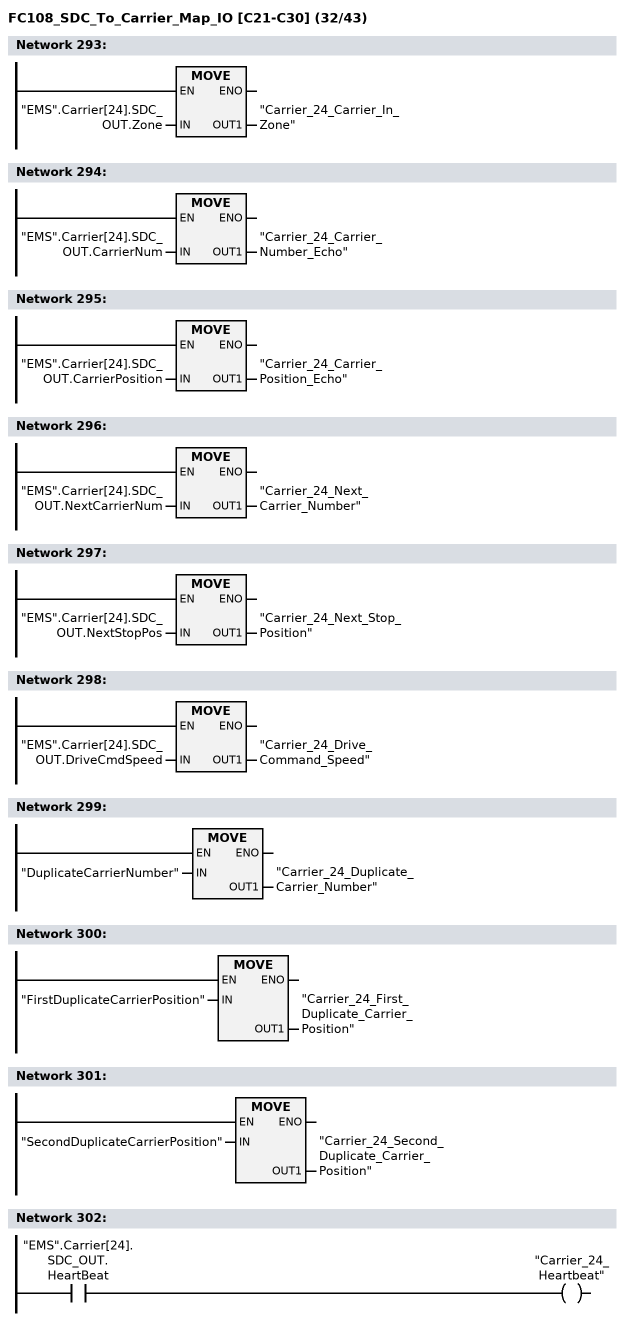
   RUNG wire#powerrail
      Move(in := "EMS".Carrier[24].SDC_OUT.Zone, out1 => "Carrier_24_Carrier_In_Zone")
   END_RUNG
   // the same network as SCL:
   "Carrier_24_Carrier_In_Zone" := "EMS".Carrier[24].SDC_OUT.Zone;
END_REGION

REGION Network 294
   RUNG wire#powerrail
      Move(in := "EMS".Carrier[24].SDC_OUT.CarrierNum, out1 => "Carrier_24_Carrier_Number_Echo")
   END_RUNG
   // the same network as SCL:
   "Carrier_24_Carrier_Number_Echo" := "EMS".Carrier[24].SDC_OUT.CarrierNum;
END_REGION

REGION Network 295
   RUNG wire#powerrail
      Move(in := "EMS".Carrier[24].SDC_OUT.CarrierPosition, out1 => "Carrier_24_Carrier_Position_Echo")
   END_RUNG
   // the same network as SCL:
   "Carrier_24_Carrier_Position_Echo" := "EMS".Carrier[24].SDC_OUT.CarrierPosition;
END_REGION

REGION Network 296
   RUNG wire#powerrail
      Move(in := "EMS".Carrier[24].SDC_OUT.NextCarrierNum, out1 => "Carrier_24_Next_Carrier_Number")
   END_RUNG
   // the same network as SCL:
   "Carrier_24_Next_Carrier_Number" := "EMS".Carrier[24].SDC_OUT.NextCarrierNum;
END_REGION

REGION Network 297
   RUNG wire#powerrail
      Move(in := "EMS".Carrier[24].SDC_OUT.NextStopPos, out1 => "Carrier_24_Next_Stop_Position")
   END_RUNG
   // the same network as SCL:
   "Carrier_24_Next_Stop_Position" := "EMS".Carrier[24].SDC_OUT.NextStopPos;
END_REGION

REGION Network 298
   RUNG wire#powerrail
      Move(in := "EMS".Carrier[24].SDC_OUT.DriveCmdSpeed, out1 => "Carrier_24_Drive_Command_Speed")
   END_RUNG
   // the same network as SCL:
   "Carrier_24_Drive_Command_Speed" := "EMS".Carrier[24].SDC_OUT.DriveCmdSpeed;
END_REGION

REGION Network 299
   RUNG wire#powerrail
      Move(in := "DuplicateCarrierNumber", out1 => "Carrier_24_Duplicate_Carrier_Number")
   END_RUNG
   // the same network as SCL:
   "Carrier_24_Duplicate_Carrier_Number" := "DuplicateCarrierNumber";
END_REGION

REGION Network 300
   RUNG wire#powerrail
      Move(in := "FirstDuplicateCarrierPosition", out1 => "Carrier_24_First_Duplicate_Carrier_Position")
   END_RUNG
   // the same network as SCL:
   "Carrier_24_First_Duplicate_Carrier_Position" := "FirstDuplicateCarrierPosition";
END_REGION

REGION Network 301
   RUNG wire#powerrail
      Move(in := "SecondDuplicateCarrierPosition", out1 => "Carrier_24_Second_Duplicate_Carrier_Position")
   END_RUNG
   // the same network as SCL:
   "Carrier_24_Second_Duplicate_Carrier_Position" := "SecondDuplicateCarrierPosition";
END_REGION

REGION Network 302
   RUNG wire#powerrail
      Contact( "EMS".Carrier[24].SDC_OUT.HeartBeat )
      Coil( "Carrier_24_Heartbeat" )
   END_RUNG
   // the same network as SCL:
   "Carrier_24_Heartbeat" := "EMS".Carrier[24].SDC_OUT.HeartBeat;
END_REGION

REGION Network 303
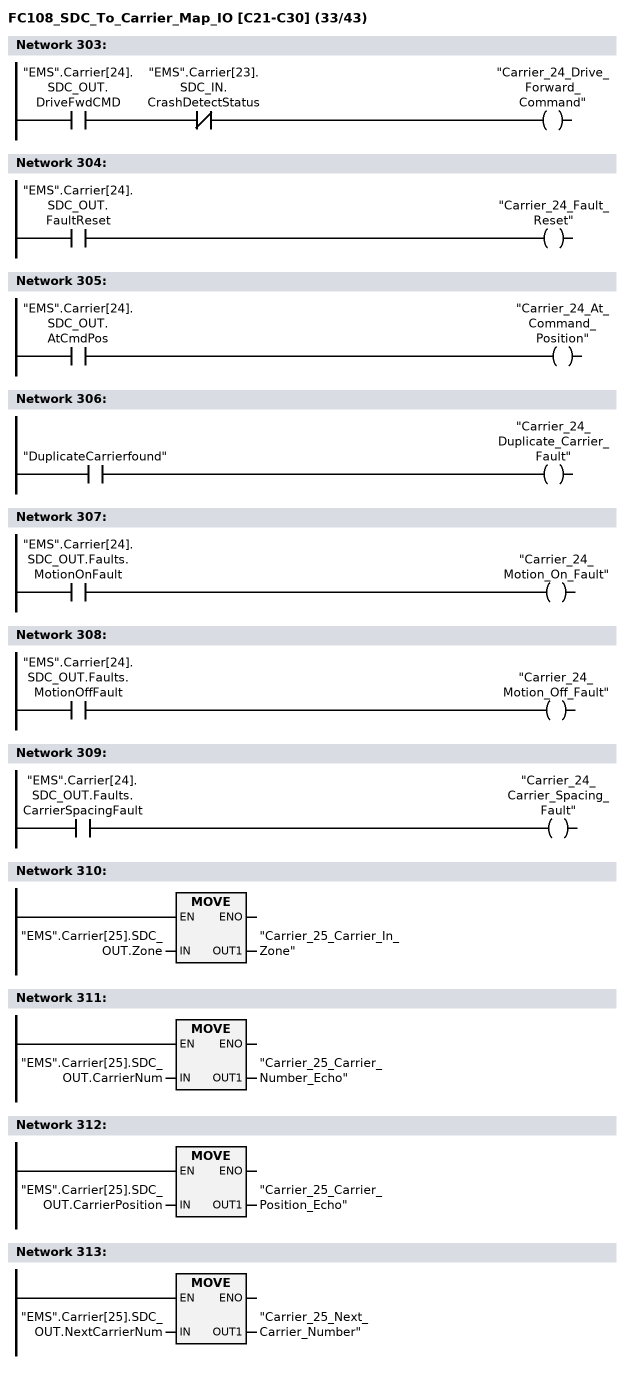
   RUNG wire#powerrail
      Contact( "EMS".Carrier[24].SDC_OUT.DriveFwdCMD )
      I_Contact( "EMS".Carrier[23].SDC_IN.CrashDetectStatus )
      Coil( "Carrier_24_Drive_Forward_Command" )
   END_RUNG
   // the same network as SCL:
   "Carrier_24_Drive_Forward_Command" := "EMS".Carrier[24].SDC_OUT.DriveFwdCMD AND NOT "EMS".Carrier[23].SDC_IN.CrashDetectStatus;
END_REGION

REGION Network 304
   RUNG wire#powerrail
      Contact( "EMS".Carrier[24].SDC_OUT.FaultReset )
      Coil( "Carrier_24_Fault_Reset" )
   END_RUNG
   // the same network as SCL:
   "Carrier_24_Fault_Reset" := "EMS".Carrier[24].SDC_OUT.FaultReset;
END_REGION

REGION Network 305
   RUNG wire#powerrail
      Contact( "EMS".Carrier[24].SDC_OUT.AtCmdPos )
      Coil( "Carrier_24_At_Command_Position" )
   END_RUNG
   // the same network as SCL:
   "Carrier_24_At_Command_Position" := "EMS".Carrier[24].SDC_OUT.AtCmdPos;
END_REGION

REGION Network 306
   RUNG wire#powerrail
      Contact( "DuplicateCarrierfound" )
      Coil( "Carrier_24_Duplicate_Carrier_Fault" )
   END_RUNG
   // the same network as SCL:
   "Carrier_24_Duplicate_Carrier_Fault" := "DuplicateCarrierfound";
END_REGION

REGION Network 307
   RUNG wire#powerrail
      Contact( "EMS".Carrier[24].SDC_OUT.Faults.MotionOnFault )
      Coil( "Carrier_24_Motion_On_Fault" )
   END_RUNG
   // the same network as SCL:
   "Carrier_24_Motion_On_Fault" := "EMS".Carrier[24].SDC_OUT.Faults.MotionOnFault;
END_REGION

REGION Network 308
   RUNG wire#powerrail
      Contact( "EMS".Carrier[24].SDC_OUT.Faults.MotionOffFault )
      Coil( "Carrier_24_Motion_Off_Fault" )
   END_RUNG
   // the same network as SCL:
   "Carrier_24_Motion_Off_Fault" := "EMS".Carrier[24].SDC_OUT.Faults.MotionOffFault;
END_REGION

REGION Network 309
   RUNG wire#powerrail
      Contact( "EMS".Carrier[24].SDC_OUT.Faults.CarrierSpacingFault )
      Coil( "Carrier_24_Carrier_Spacing_Fault" )
   END_RUNG
   // the same network as SCL:
   "Carrier_24_Carrier_Spacing_Fault" := "EMS".Carrier[24].SDC_OUT.Faults.CarrierSpacingFault;
END_REGION

REGION Network 310
   RUNG wire#powerrail
      Move(in := "EMS".Carrier[25].SDC_OUT.Zone, out1 => "Carrier_25_Carrier_In_Zone")
   END_RUNG
   // the same network as SCL:
   "Carrier_25_Carrier_In_Zone" := "EMS".Carrier[25].SDC_OUT.Zone;
END_REGION

REGION Network 311
   RUNG wire#powerrail
      Move(in := "EMS".Carrier[25].SDC_OUT.CarrierNum, out1 => "Carrier_25_Carrier_Number_Echo")
   END_RUNG
   // the same network as SCL:
   "Carrier_25_Carrier_Number_Echo" := "EMS".Carrier[25].SDC_OUT.CarrierNum;
END_REGION

REGION Network 312
   RUNG wire#powerrail
      Move(in := "EMS".Carrier[25].SDC_OUT.CarrierPosition, out1 => "Carrier_25_Carrier_Position_Echo")
   END_RUNG
   // the same network as SCL:
   "Carrier_25_Carrier_Position_Echo" := "EMS".Carrier[25].SDC_OUT.CarrierPosition;
END_REGION

REGION Network 313
   RUNG wire#powerrail
      Move(in := "EMS".Carrier[25].SDC_OUT.NextCarrierNum, out1 => "Carrier_25_Next_Carrier_Number")
   END_RUNG
   // the same network as SCL:
   "Carrier_25_Next_Carrier_Number" := "EMS".Carrier[25].SDC_OUT.NextCarrierNum;
END_REGION

REGION Network 314
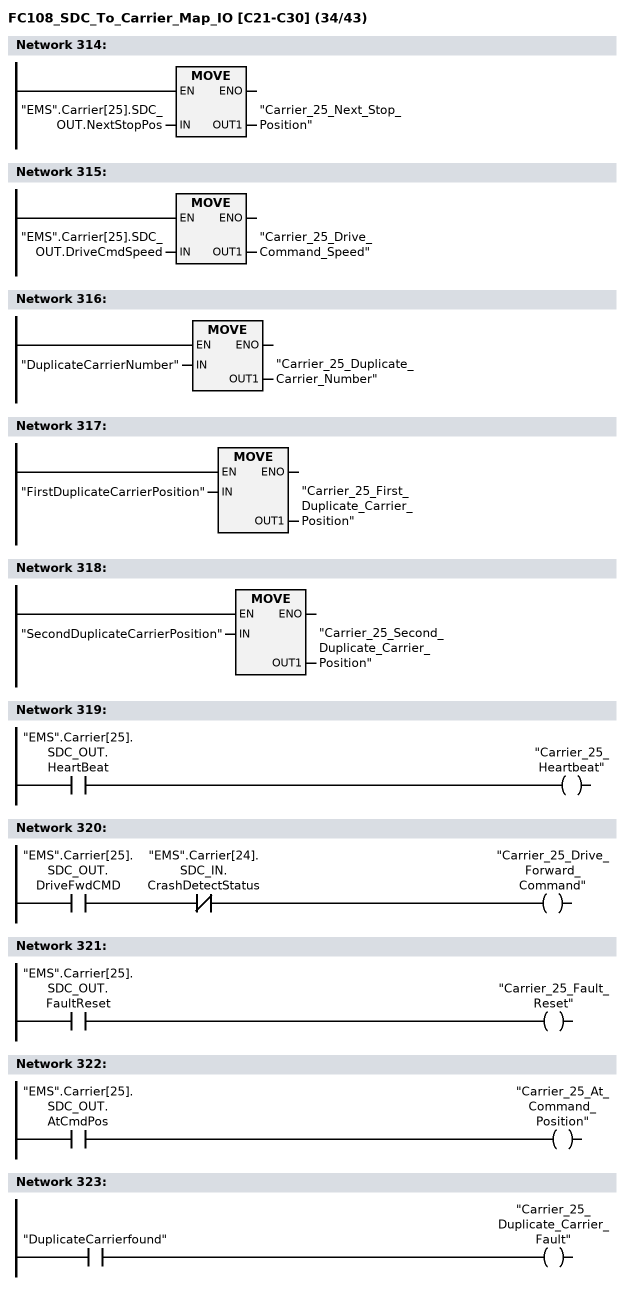
   RUNG wire#powerrail
      Move(in := "EMS".Carrier[25].SDC_OUT.NextStopPos, out1 => "Carrier_25_Next_Stop_Position")
   END_RUNG
   // the same network as SCL:
   "Carrier_25_Next_Stop_Position" := "EMS".Carrier[25].SDC_OUT.NextStopPos;
END_REGION

REGION Network 315
   RUNG wire#powerrail
      Move(in := "EMS".Carrier[25].SDC_OUT.DriveCmdSpeed, out1 => "Carrier_25_Drive_Command_Speed")
   END_RUNG
   // the same network as SCL:
   "Carrier_25_Drive_Command_Speed" := "EMS".Carrier[25].SDC_OUT.DriveCmdSpeed;
END_REGION

REGION Network 316
   RUNG wire#powerrail
      Move(in := "DuplicateCarrierNumber", out1 => "Carrier_25_Duplicate_Carrier_Number")
   END_RUNG
   // the same network as SCL:
   "Carrier_25_Duplicate_Carrier_Number" := "DuplicateCarrierNumber";
END_REGION

REGION Network 317
   RUNG wire#powerrail
      Move(in := "FirstDuplicateCarrierPosition", out1 => "Carrier_25_First_Duplicate_Carrier_Position")
   END_RUNG
   // the same network as SCL:
   "Carrier_25_First_Duplicate_Carrier_Position" := "FirstDuplicateCarrierPosition";
END_REGION

REGION Network 318
   RUNG wire#powerrail
      Move(in := "SecondDuplicateCarrierPosition", out1 => "Carrier_25_Second_Duplicate_Carrier_Position")
   END_RUNG
   // the same network as SCL:
   "Carrier_25_Second_Duplicate_Carrier_Position" := "SecondDuplicateCarrierPosition";
END_REGION

REGION Network 319
   RUNG wire#powerrail
      Contact( "EMS".Carrier[25].SDC_OUT.HeartBeat )
      Coil( "Carrier_25_Heartbeat" )
   END_RUNG
   // the same network as SCL:
   "Carrier_25_Heartbeat" := "EMS".Carrier[25].SDC_OUT.HeartBeat;
END_REGION

REGION Network 320
   RUNG wire#powerrail
      Contact( "EMS".Carrier[25].SDC_OUT.DriveFwdCMD )
      I_Contact( "EMS".Carrier[24].SDC_IN.CrashDetectStatus )
      Coil( "Carrier_25_Drive_Forward_Command" )
   END_RUNG
   // the same network as SCL:
   "Carrier_25_Drive_Forward_Command" := "EMS".Carrier[25].SDC_OUT.DriveFwdCMD AND NOT "EMS".Carrier[24].SDC_IN.CrashDetectStatus;
END_REGION

REGION Network 321
   RUNG wire#powerrail
      Contact( "EMS".Carrier[25].SDC_OUT.FaultReset )
      Coil( "Carrier_25_Fault_Reset" )
   END_RUNG
   // the same network as SCL:
   "Carrier_25_Fault_Reset" := "EMS".Carrier[25].SDC_OUT.FaultReset;
END_REGION

REGION Network 322
   RUNG wire#powerrail
      Contact( "EMS".Carrier[25].SDC_OUT.AtCmdPos )
      Coil( "Carrier_25_At_Command_Position" )
   END_RUNG
   // the same network as SCL:
   "Carrier_25_At_Command_Position" := "EMS".Carrier[25].SDC_OUT.AtCmdPos;
END_REGION

REGION Network 323
   RUNG wire#powerrail
      Contact( "DuplicateCarrierfound" )
      Coil( "Carrier_25_Duplicate_Carrier_Fault" )
   END_RUNG
   // the same network as SCL:
   "Carrier_25_Duplicate_Carrier_Fault" := "DuplicateCarrierfound";
END_REGION

REGION Network 324
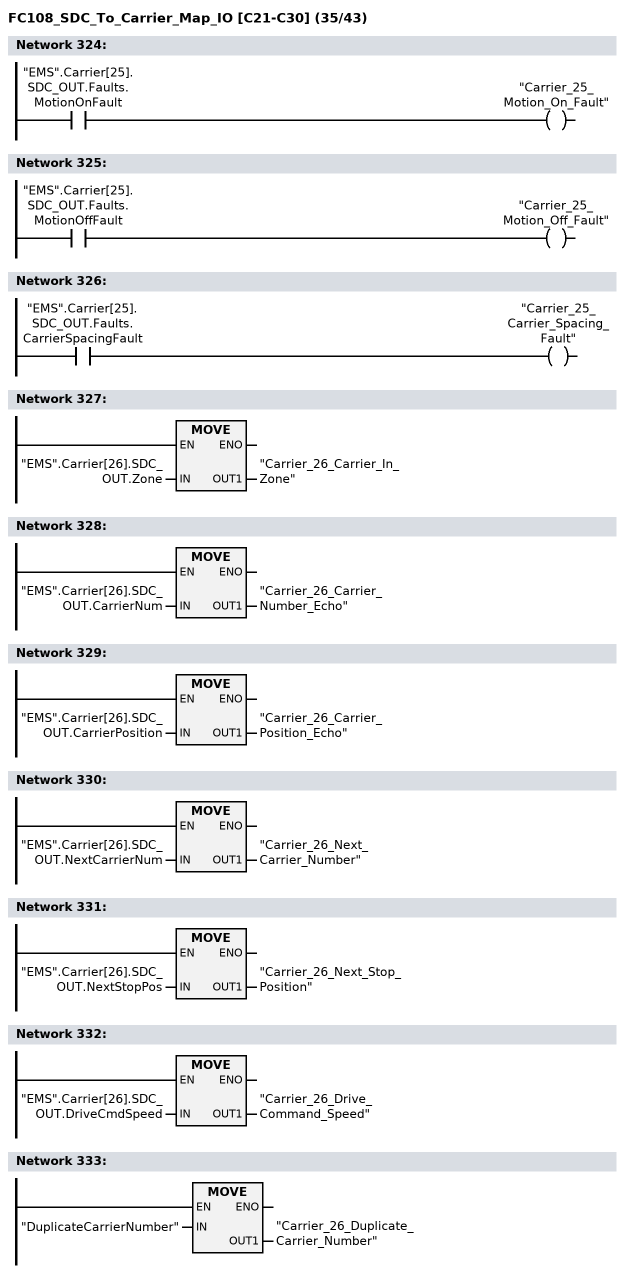
   RUNG wire#powerrail
      Contact( "EMS".Carrier[25].SDC_OUT.Faults.MotionOnFault )
      Coil( "Carrier_25_Motion_On_Fault" )
   END_RUNG
   // the same network as SCL:
   "Carrier_25_Motion_On_Fault" := "EMS".Carrier[25].SDC_OUT.Faults.MotionOnFault;
END_REGION

REGION Network 325
   RUNG wire#powerrail
      Contact( "EMS".Carrier[25].SDC_OUT.Faults.MotionOffFault )
      Coil( "Carrier_25_Motion_Off_Fault" )
   END_RUNG
   // the same network as SCL:
   "Carrier_25_Motion_Off_Fault" := "EMS".Carrier[25].SDC_OUT.Faults.MotionOffFault;
END_REGION

REGION Network 326
   RUNG wire#powerrail
      Contact( "EMS".Carrier[25].SDC_OUT.Faults.CarrierSpacingFault )
      Coil( "Carrier_25_Carrier_Spacing_Fault" )
   END_RUNG
   // the same network as SCL:
   "Carrier_25_Carrier_Spacing_Fault" := "EMS".Carrier[25].SDC_OUT.Faults.CarrierSpacingFault;
END_REGION

REGION Network 327
   RUNG wire#powerrail
      Move(in := "EMS".Carrier[26].SDC_OUT.Zone, out1 => "Carrier_26_Carrier_In_Zone")
   END_RUNG
   // the same network as SCL:
   "Carrier_26_Carrier_In_Zone" := "EMS".Carrier[26].SDC_OUT.Zone;
END_REGION

REGION Network 328
   RUNG wire#powerrail
      Move(in := "EMS".Carrier[26].SDC_OUT.CarrierNum, out1 => "Carrier_26_Carrier_Number_Echo")
   END_RUNG
   // the same network as SCL:
   "Carrier_26_Carrier_Number_Echo" := "EMS".Carrier[26].SDC_OUT.CarrierNum;
END_REGION

REGION Network 329
   RUNG wire#powerrail
      Move(in := "EMS".Carrier[26].SDC_OUT.CarrierPosition, out1 => "Carrier_26_Carrier_Position_Echo")
   END_RUNG
   // the same network as SCL:
   "Carrier_26_Carrier_Position_Echo" := "EMS".Carrier[26].SDC_OUT.CarrierPosition;
END_REGION

REGION Network 330
   RUNG wire#powerrail
      Move(in := "EMS".Carrier[26].SDC_OUT.NextCarrierNum, out1 => "Carrier_26_Next_Carrier_Number")
   END_RUNG
   // the same network as SCL:
   "Carrier_26_Next_Carrier_Number" := "EMS".Carrier[26].SDC_OUT.NextCarrierNum;
END_REGION

REGION Network 331
   RUNG wire#powerrail
      Move(in := "EMS".Carrier[26].SDC_OUT.NextStopPos, out1 => "Carrier_26_Next_Stop_Position")
   END_RUNG
   // the same network as SCL:
   "Carrier_26_Next_Stop_Position" := "EMS".Carrier[26].SDC_OUT.NextStopPos;
END_REGION

REGION Network 332
   RUNG wire#powerrail
      Move(in := "EMS".Carrier[26].SDC_OUT.DriveCmdSpeed, out1 => "Carrier_26_Drive_Command_Speed")
   END_RUNG
   // the same network as SCL:
   "Carrier_26_Drive_Command_Speed" := "EMS".Carrier[26].SDC_OUT.DriveCmdSpeed;
END_REGION

REGION Network 333
   RUNG wire#powerrail
      Move(in := "DuplicateCarrierNumber", out1 => "Carrier_26_Duplicate_Carrier_Number")
   END_RUNG
   // the same network as SCL:
   "Carrier_26_Duplicate_Carrier_Number" := "DuplicateCarrierNumber";
END_REGION

REGION Network 334
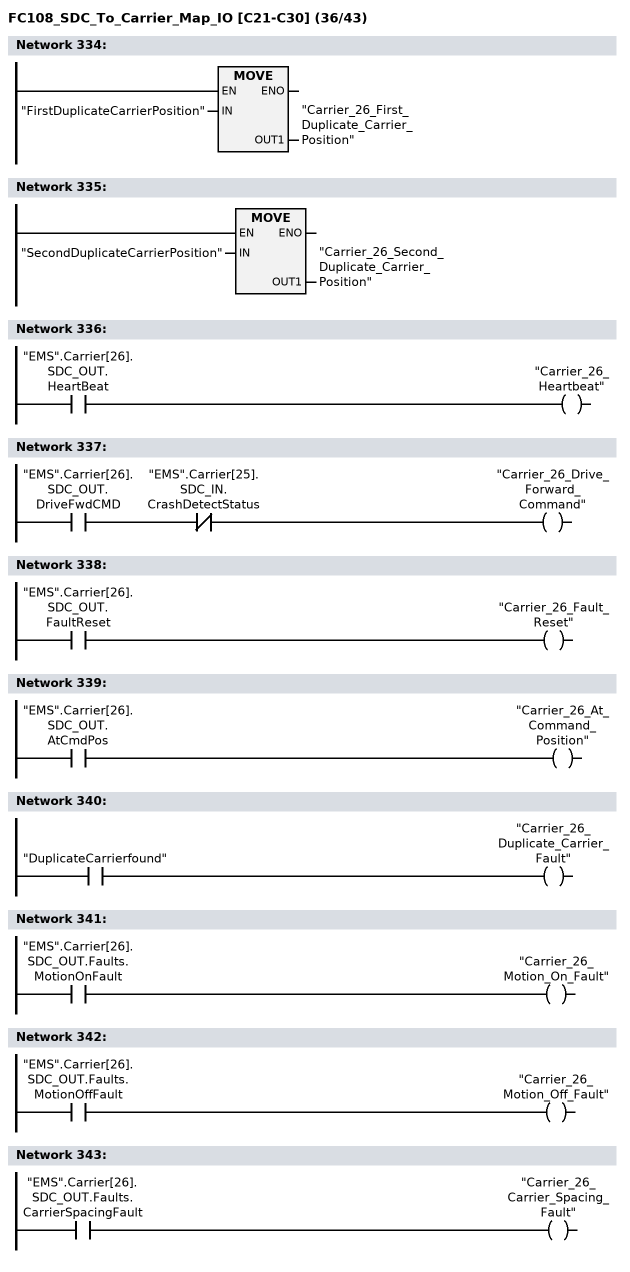
   RUNG wire#powerrail
      Move(in := "FirstDuplicateCarrierPosition", out1 => "Carrier_26_First_Duplicate_Carrier_Position")
   END_RUNG
   // the same network as SCL:
   "Carrier_26_First_Duplicate_Carrier_Position" := "FirstDuplicateCarrierPosition";
END_REGION

REGION Network 335
   RUNG wire#powerrail
      Move(in := "SecondDuplicateCarrierPosition", out1 => "Carrier_26_Second_Duplicate_Carrier_Position")
   END_RUNG
   // the same network as SCL:
   "Carrier_26_Second_Duplicate_Carrier_Position" := "SecondDuplicateCarrierPosition";
END_REGION

REGION Network 336
   RUNG wire#powerrail
      Contact( "EMS".Carrier[26].SDC_OUT.HeartBeat )
      Coil( "Carrier_26_Heartbeat" )
   END_RUNG
   // the same network as SCL:
   "Carrier_26_Heartbeat" := "EMS".Carrier[26].SDC_OUT.HeartBeat;
END_REGION

REGION Network 337
   RUNG wire#powerrail
      Contact( "EMS".Carrier[26].SDC_OUT.DriveFwdCMD )
      I_Contact( "EMS".Carrier[25].SDC_IN.CrashDetectStatus )
      Coil( "Carrier_26_Drive_Forward_Command" )
   END_RUNG
   // the same network as SCL:
   "Carrier_26_Drive_Forward_Command" := "EMS".Carrier[26].SDC_OUT.DriveFwdCMD AND NOT "EMS".Carrier[25].SDC_IN.CrashDetectStatus;
END_REGION

REGION Network 338
   RUNG wire#powerrail
      Contact( "EMS".Carrier[26].SDC_OUT.FaultReset )
      Coil( "Carrier_26_Fault_Reset" )
   END_RUNG
   // the same network as SCL:
   "Carrier_26_Fault_Reset" := "EMS".Carrier[26].SDC_OUT.FaultReset;
END_REGION

REGION Network 339
   RUNG wire#powerrail
      Contact( "EMS".Carrier[26].SDC_OUT.AtCmdPos )
      Coil( "Carrier_26_At_Command_Position" )
   END_RUNG
   // the same network as SCL:
   "Carrier_26_At_Command_Position" := "EMS".Carrier[26].SDC_OUT.AtCmdPos;
END_REGION

REGION Network 340
   RUNG wire#powerrail
      Contact( "DuplicateCarrierfound" )
      Coil( "Carrier_26_Duplicate_Carrier_Fault" )
   END_RUNG
   // the same network as SCL:
   "Carrier_26_Duplicate_Carrier_Fault" := "DuplicateCarrierfound";
END_REGION

REGION Network 341
   RUNG wire#powerrail
      Contact( "EMS".Carrier[26].SDC_OUT.Faults.MotionOnFault )
      Coil( "Carrier_26_Motion_On_Fault" )
   END_RUNG
   // the same network as SCL:
   "Carrier_26_Motion_On_Fault" := "EMS".Carrier[26].SDC_OUT.Faults.MotionOnFault;
END_REGION

REGION Network 342
   RUNG wire#powerrail
      Contact( "EMS".Carrier[26].SDC_OUT.Faults.MotionOffFault )
      Coil( "Carrier_26_Motion_Off_Fault" )
   END_RUNG
   // the same network as SCL:
   "Carrier_26_Motion_Off_Fault" := "EMS".Carrier[26].SDC_OUT.Faults.MotionOffFault;
END_REGION

REGION Network 343
   RUNG wire#powerrail
      Contact( "EMS".Carrier[26].SDC_OUT.Faults.CarrierSpacingFault )
      Coil( "Carrier_26_Carrier_Spacing_Fault" )
   END_RUNG
   // the same network as SCL:
   "Carrier_26_Carrier_Spacing_Fault" := "EMS".Carrier[26].SDC_OUT.Faults.CarrierSpacingFault;
END_REGION

REGION Network 344
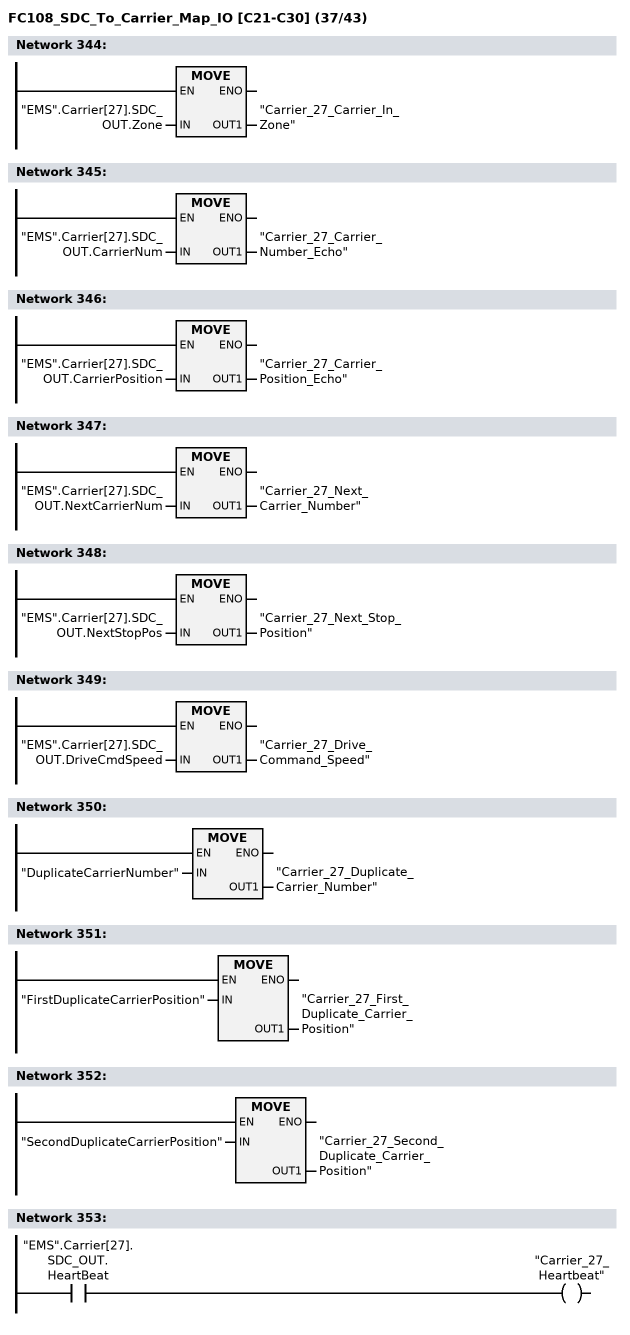
   RUNG wire#powerrail
      Move(in := "EMS".Carrier[27].SDC_OUT.Zone, out1 => "Carrier_27_Carrier_In_Zone")
   END_RUNG
   // the same network as SCL:
   "Carrier_27_Carrier_In_Zone" := "EMS".Carrier[27].SDC_OUT.Zone;
END_REGION

REGION Network 345
   RUNG wire#powerrail
      Move(in := "EMS".Carrier[27].SDC_OUT.CarrierNum, out1 => "Carrier_27_Carrier_Number_Echo")
   END_RUNG
   // the same network as SCL:
   "Carrier_27_Carrier_Number_Echo" := "EMS".Carrier[27].SDC_OUT.CarrierNum;
END_REGION

REGION Network 346
   RUNG wire#powerrail
      Move(in := "EMS".Carrier[27].SDC_OUT.CarrierPosition, out1 => "Carrier_27_Carrier_Position_Echo")
   END_RUNG
   // the same network as SCL:
   "Carrier_27_Carrier_Position_Echo" := "EMS".Carrier[27].SDC_OUT.CarrierPosition;
END_REGION

REGION Network 347
   RUNG wire#powerrail
      Move(in := "EMS".Carrier[27].SDC_OUT.NextCarrierNum, out1 => "Carrier_27_Next_Carrier_Number")
   END_RUNG
   // the same network as SCL:
   "Carrier_27_Next_Carrier_Number" := "EMS".Carrier[27].SDC_OUT.NextCarrierNum;
END_REGION

REGION Network 348
   RUNG wire#powerrail
      Move(in := "EMS".Carrier[27].SDC_OUT.NextStopPos, out1 => "Carrier_27_Next_Stop_Position")
   END_RUNG
   // the same network as SCL:
   "Carrier_27_Next_Stop_Position" := "EMS".Carrier[27].SDC_OUT.NextStopPos;
END_REGION

REGION Network 349
   RUNG wire#powerrail
      Move(in := "EMS".Carrier[27].SDC_OUT.DriveCmdSpeed, out1 => "Carrier_27_Drive_Command_Speed")
   END_RUNG
   // the same network as SCL:
   "Carrier_27_Drive_Command_Speed" := "EMS".Carrier[27].SDC_OUT.DriveCmdSpeed;
END_REGION

REGION Network 350
   RUNG wire#powerrail
      Move(in := "DuplicateCarrierNumber", out1 => "Carrier_27_Duplicate_Carrier_Number")
   END_RUNG
   // the same network as SCL:
   "Carrier_27_Duplicate_Carrier_Number" := "DuplicateCarrierNumber";
END_REGION

REGION Network 351
   RUNG wire#powerrail
      Move(in := "FirstDuplicateCarrierPosition", out1 => "Carrier_27_First_Duplicate_Carrier_Position")
   END_RUNG
   // the same network as SCL:
   "Carrier_27_First_Duplicate_Carrier_Position" := "FirstDuplicateCarrierPosition";
END_REGION

REGION Network 352
   RUNG wire#powerrail
      Move(in := "SecondDuplicateCarrierPosition", out1 => "Carrier_27_Second_Duplicate_Carrier_Position")
   END_RUNG
   // the same network as SCL:
   "Carrier_27_Second_Duplicate_Carrier_Position" := "SecondDuplicateCarrierPosition";
END_REGION

REGION Network 353
   RUNG wire#powerrail
      Contact( "EMS".Carrier[27].SDC_OUT.HeartBeat )
      Coil( "Carrier_27_Heartbeat" )
   END_RUNG
   // the same network as SCL:
   "Carrier_27_Heartbeat" := "EMS".Carrier[27].SDC_OUT.HeartBeat;
END_REGION

REGION Network 354
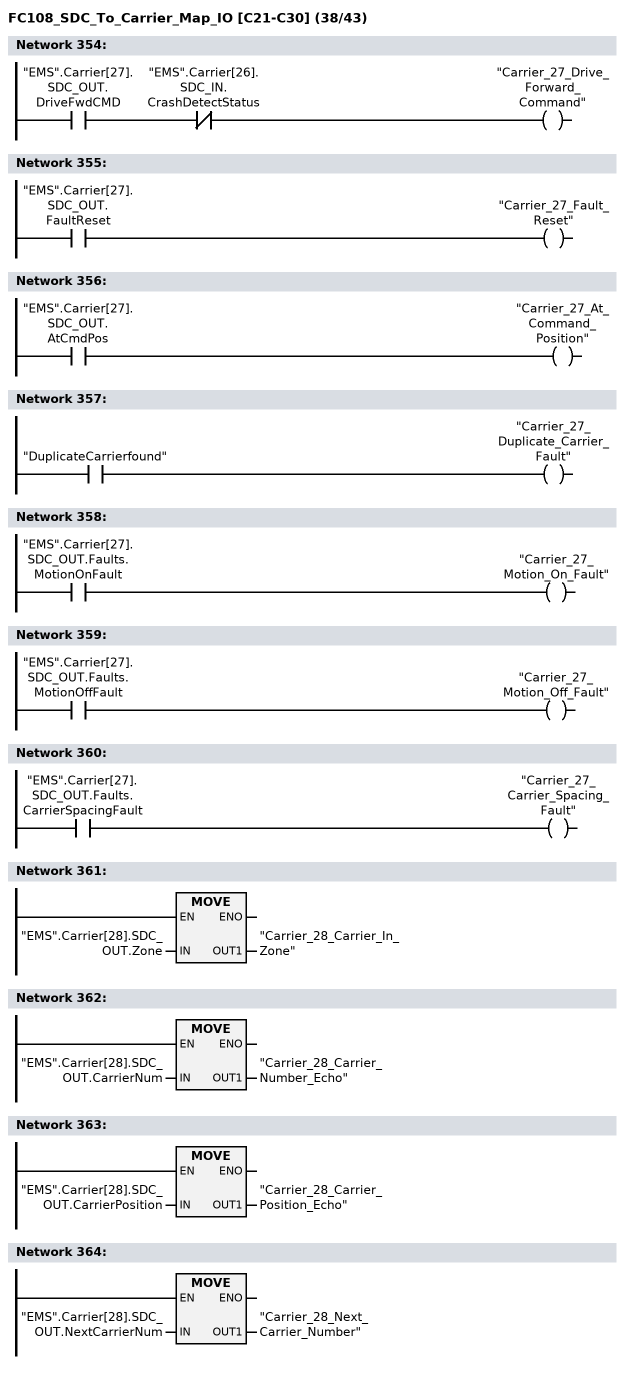
   RUNG wire#powerrail
      Contact( "EMS".Carrier[27].SDC_OUT.DriveFwdCMD )
      I_Contact( "EMS".Carrier[26].SDC_IN.CrashDetectStatus )
      Coil( "Carrier_27_Drive_Forward_Command" )
   END_RUNG
   // the same network as SCL:
   "Carrier_27_Drive_Forward_Command" := "EMS".Carrier[27].SDC_OUT.DriveFwdCMD AND NOT "EMS".Carrier[26].SDC_IN.CrashDetectStatus;
END_REGION

REGION Network 355
   RUNG wire#powerrail
      Contact( "EMS".Carrier[27].SDC_OUT.FaultReset )
      Coil( "Carrier_27_Fault_Reset" )
   END_RUNG
   // the same network as SCL:
   "Carrier_27_Fault_Reset" := "EMS".Carrier[27].SDC_OUT.FaultReset;
END_REGION

REGION Network 356
   RUNG wire#powerrail
      Contact( "EMS".Carrier[27].SDC_OUT.AtCmdPos )
      Coil( "Carrier_27_At_Command_Position" )
   END_RUNG
   // the same network as SCL:
   "Carrier_27_At_Command_Position" := "EMS".Carrier[27].SDC_OUT.AtCmdPos;
END_REGION

REGION Network 357
   RUNG wire#powerrail
      Contact( "DuplicateCarrierfound" )
      Coil( "Carrier_27_Duplicate_Carrier_Fault" )
   END_RUNG
   // the same network as SCL:
   "Carrier_27_Duplicate_Carrier_Fault" := "DuplicateCarrierfound";
END_REGION

REGION Network 358
   RUNG wire#powerrail
      Contact( "EMS".Carrier[27].SDC_OUT.Faults.MotionOnFault )
      Coil( "Carrier_27_Motion_On_Fault" )
   END_RUNG
   // the same network as SCL:
   "Carrier_27_Motion_On_Fault" := "EMS".Carrier[27].SDC_OUT.Faults.MotionOnFault;
END_REGION

REGION Network 359
   RUNG wire#powerrail
      Contact( "EMS".Carrier[27].SDC_OUT.Faults.MotionOffFault )
      Coil( "Carrier_27_Motion_Off_Fault" )
   END_RUNG
   // the same network as SCL:
   "Carrier_27_Motion_Off_Fault" := "EMS".Carrier[27].SDC_OUT.Faults.MotionOffFault;
END_REGION

REGION Network 360
   RUNG wire#powerrail
      Contact( "EMS".Carrier[27].SDC_OUT.Faults.CarrierSpacingFault )
      Coil( "Carrier_27_Carrier_Spacing_Fault" )
   END_RUNG
   // the same network as SCL:
   "Carrier_27_Carrier_Spacing_Fault" := "EMS".Carrier[27].SDC_OUT.Faults.CarrierSpacingFault;
END_REGION

REGION Network 361
   RUNG wire#powerrail
      Move(in := "EMS".Carrier[28].SDC_OUT.Zone, out1 => "Carrier_28_Carrier_In_Zone")
   END_RUNG
   // the same network as SCL:
   "Carrier_28_Carrier_In_Zone" := "EMS".Carrier[28].SDC_OUT.Zone;
END_REGION

REGION Network 362
   RUNG wire#powerrail
      Move(in := "EMS".Carrier[28].SDC_OUT.CarrierNum, out1 => "Carrier_28_Carrier_Number_Echo")
   END_RUNG
   // the same network as SCL:
   "Carrier_28_Carrier_Number_Echo" := "EMS".Carrier[28].SDC_OUT.CarrierNum;
END_REGION

REGION Network 363
   RUNG wire#powerrail
      Move(in := "EMS".Carrier[28].SDC_OUT.CarrierPosition, out1 => "Carrier_28_Carrier_Position_Echo")
   END_RUNG
   // the same network as SCL:
   "Carrier_28_Carrier_Position_Echo" := "EMS".Carrier[28].SDC_OUT.CarrierPosition;
END_REGION

REGION Network 364
   RUNG wire#powerrail
      Move(in := "EMS".Carrier[28].SDC_OUT.NextCarrierNum, out1 => "Carrier_28_Next_Carrier_Number")
   END_RUNG
   // the same network as SCL:
   "Carrier_28_Next_Carrier_Number" := "EMS".Carrier[28].SDC_OUT.NextCarrierNum;
END_REGION

REGION Network 365
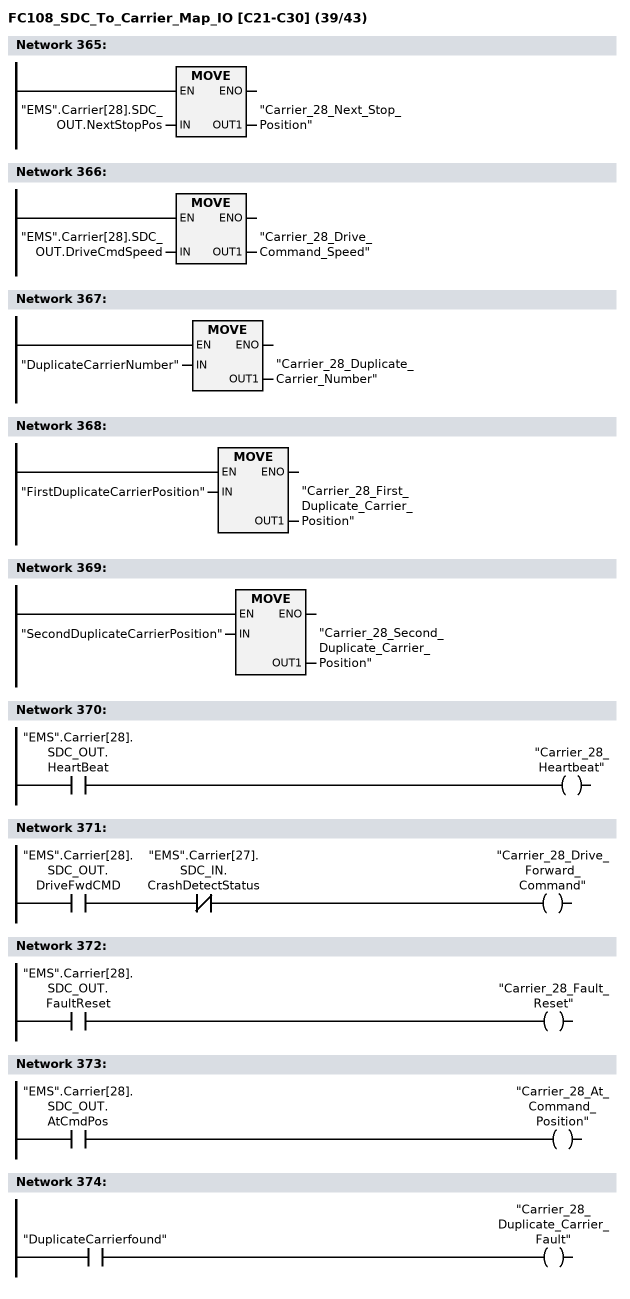
   RUNG wire#powerrail
      Move(in := "EMS".Carrier[28].SDC_OUT.NextStopPos, out1 => "Carrier_28_Next_Stop_Position")
   END_RUNG
   // the same network as SCL:
   "Carrier_28_Next_Stop_Position" := "EMS".Carrier[28].SDC_OUT.NextStopPos;
END_REGION

REGION Network 366
   RUNG wire#powerrail
      Move(in := "EMS".Carrier[28].SDC_OUT.DriveCmdSpeed, out1 => "Carrier_28_Drive_Command_Speed")
   END_RUNG
   // the same network as SCL:
   "Carrier_28_Drive_Command_Speed" := "EMS".Carrier[28].SDC_OUT.DriveCmdSpeed;
END_REGION

REGION Network 367
   RUNG wire#powerrail
      Move(in := "DuplicateCarrierNumber", out1 => "Carrier_28_Duplicate_Carrier_Number")
   END_RUNG
   // the same network as SCL:
   "Carrier_28_Duplicate_Carrier_Number" := "DuplicateCarrierNumber";
END_REGION

REGION Network 368
   RUNG wire#powerrail
      Move(in := "FirstDuplicateCarrierPosition", out1 => "Carrier_28_First_Duplicate_Carrier_Position")
   END_RUNG
   // the same network as SCL:
   "Carrier_28_First_Duplicate_Carrier_Position" := "FirstDuplicateCarrierPosition";
END_REGION

REGION Network 369
   RUNG wire#powerrail
      Move(in := "SecondDuplicateCarrierPosition", out1 => "Carrier_28_Second_Duplicate_Carrier_Position")
   END_RUNG
   // the same network as SCL:
   "Carrier_28_Second_Duplicate_Carrier_Position" := "SecondDuplicateCarrierPosition";
END_REGION

REGION Network 370
   RUNG wire#powerrail
      Contact( "EMS".Carrier[28].SDC_OUT.HeartBeat )
      Coil( "Carrier_28_Heartbeat" )
   END_RUNG
   // the same network as SCL:
   "Carrier_28_Heartbeat" := "EMS".Carrier[28].SDC_OUT.HeartBeat;
END_REGION

REGION Network 371
   RUNG wire#powerrail
      Contact( "EMS".Carrier[28].SDC_OUT.DriveFwdCMD )
      I_Contact( "EMS".Carrier[27].SDC_IN.CrashDetectStatus )
      Coil( "Carrier_28_Drive_Forward_Command" )
   END_RUNG
   // the same network as SCL:
   "Carrier_28_Drive_Forward_Command" := "EMS".Carrier[28].SDC_OUT.DriveFwdCMD AND NOT "EMS".Carrier[27].SDC_IN.CrashDetectStatus;
END_REGION

REGION Network 372
   RUNG wire#powerrail
      Contact( "EMS".Carrier[28].SDC_OUT.FaultReset )
      Coil( "Carrier_28_Fault_Reset" )
   END_RUNG
   // the same network as SCL:
   "Carrier_28_Fault_Reset" := "EMS".Carrier[28].SDC_OUT.FaultReset;
END_REGION

REGION Network 373
   RUNG wire#powerrail
      Contact( "EMS".Carrier[28].SDC_OUT.AtCmdPos )
      Coil( "Carrier_28_At_Command_Position" )
   END_RUNG
   // the same network as SCL:
   "Carrier_28_At_Command_Position" := "EMS".Carrier[28].SDC_OUT.AtCmdPos;
END_REGION

REGION Network 374
   RUNG wire#powerrail
      Contact( "DuplicateCarrierfound" )
      Coil( "Carrier_28_Duplicate_Carrier_Fault" )
   END_RUNG
   // the same network as SCL:
   "Carrier_28_Duplicate_Carrier_Fault" := "DuplicateCarrierfound";
END_REGION

REGION Network 375
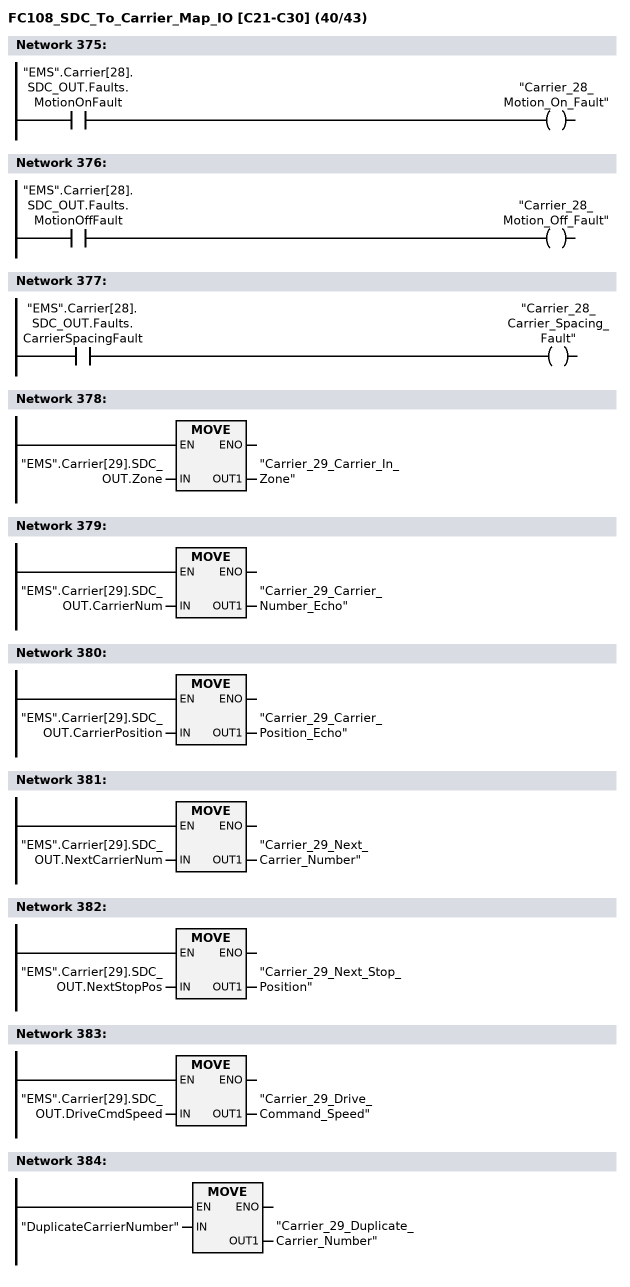
   RUNG wire#powerrail
      Contact( "EMS".Carrier[28].SDC_OUT.Faults.MotionOnFault )
      Coil( "Carrier_28_Motion_On_Fault" )
   END_RUNG
   // the same network as SCL:
   "Carrier_28_Motion_On_Fault" := "EMS".Carrier[28].SDC_OUT.Faults.MotionOnFault;
END_REGION

REGION Network 376
   RUNG wire#powerrail
      Contact( "EMS".Carrier[28].SDC_OUT.Faults.MotionOffFault )
      Coil( "Carrier_28_Motion_Off_Fault" )
   END_RUNG
   // the same network as SCL:
   "Carrier_28_Motion_Off_Fault" := "EMS".Carrier[28].SDC_OUT.Faults.MotionOffFault;
END_REGION

REGION Network 377
   RUNG wire#powerrail
      Contact( "EMS".Carrier[28].SDC_OUT.Faults.CarrierSpacingFault )
      Coil( "Carrier_28_Carrier_Spacing_Fault" )
   END_RUNG
   // the same network as SCL:
   "Carrier_28_Carrier_Spacing_Fault" := "EMS".Carrier[28].SDC_OUT.Faults.CarrierSpacingFault;
END_REGION
